(* Logix 5000 project; controller PLC_MCC1300_75F1 vendor 1 type 14 code 166 rev 32.11; software revision 32.04; part 68 of 83 *)
(* tags used below, declared in another part *)
   CM_AreaStackerToLine_JS1_Sync : CM_AreaStackerToLine;
   CM_ConveyorStackerToLine_JS1_Sync : CM_ConveyorStackerToLine;
   CM_DATA_Z410_Rx_Sync : UDT_PlateData_Convoy;
   CM_DATA_Z410_Tx : UDT_PlateData_Convoy;
   CM_DATA_Z410_Tx_PH : DINT;
   CM_LineToAreaStacker_JS1 : CM_LineToAreaStacker;
   CM_LineToConveyorStacker_JS1 : CM_LineToConveyorStacker;
   CM_LineToConveyorStacker_JS2 : CM_LineToConveyorStacker;
   GP_AccessArea_M311S_STC : GP_AccessArea_STC;
   GP_ConvertDataFromStacker : GP_ConvertDataFromStacker;
   GP_ConvertDataToStacker : GP_ConvertDataToStacker;
   Gp_SpaceConvUtilities_V1 : GP_SpaceConvUtilities_V1;
   M311 : MAC_Conveyor;
   M311_SpaceConv_Utilities : SpaceConv_Utilities;
   M316 : MAC_Conveyor;
   M316_SpaceConv_Utilities : SpaceConv_Utilities;
   M317 : MAC_Conveyor_Single;
   M317_Data : UDT_Convoy_SL;
   M317_dTractionRecovery_M3 : DINT;
   M317_dTractionRecovery_M4 : DINT;
   M317_HMR : MAC_Conveyor_HMR;
   M317_HMW : MAC_Conveyor_HMW;
   M317_M3_DR_IN_MAM : MOTION_INSTRUCTION;
   M317_M3_DR_IN_MRP : MOTION_INSTRUCTION;
   M317_SpaceConv_Utilities : SpaceConv_Utilities;
   M317_xEnableTractionRecovering : BOOL;
   M317_xLateralTractionRecovered : BOOL;
   M317_xSendCulletReqActive : BOOL;
   O : INT[128];
   TMP_CenterLites : BOOL;
   TMP_d : DINT;
   TMP_dDecelerationPositionEndConveyor : DINT;
   TMP_DistanceLateralSquaringToCenter : DINT;
   TMP_dOffsetLoadUnload_cmm : DINT;
   TMP_SendToCullet : BOOL;
   TMP_SquaringPosition : DINT;
   TMP_xConveyorOfStartCleaning : BOOL;
   TMP_xCulletPresent : BOOL;
   TMP_xLiteThisDestPresent : BOOL;
   xAlwaysOFF : BOOL;
   xAlwaysON : BOOL;
   xDebugOFF : BOOL;
   Z402 : MAC_Zone;
   Z402_HMR : MAC_Zone_HMR;
   Z402S_INPUT_xSafetyAreaPopup : BOOL;
(* MainProgram, continued *)

   // Calculation Space for Wait Stop Next Conveyor
   39: CPT(TMP_dDecelerationPositionEndConveyor,M317_SpaceConv_Utilities.CONST_dConveyorLength_cmm - M317.AUX_dAccSpace_cmm + 1000);
   // Wait stop next Machine
   40: XIO(M317.PH_x.8)GEQ(M317_SpaceConv_Utilities.O_dHeadPosition_cmm,TMP_dDecelerationPositionEndConveyor)OTE(M317.ST_xWaitStopNextMachine);
   // Set Wait Machine Stop
   41: [XIC(M317.PH_x.7) [XIO(xAlwaysOFF) ,XIC(M317.ST_xWaitStopNextMachine) [XIC(M311_SpaceConv_Utilities.O_xRampInProgress) ,XIO(M311_SpaceConv_Utilities.ST_xFeedbackRotation) ] ] ,XIC(M317.PH_x.0) NEQ(Z402_HMR.dLineSpeed_mm_min,M317.AUX_dReqSpeed_mm_min) ]OTL(M317.ST_xWaitMachineStop);
   // Reset Wait Machine Stop
   42: XIO(M317_SpaceConv_Utilities.ST_xFeedbackRotation)[XIO(M317_SpaceConv_Utilities.ST_xFeedbackRotation) ,XIO(M317.ST_xWaitStopNextMachine) ]EQU(Z402_HMR.dLineSpeed_mm_min,M317.AUX_dReqSpeed_mm_min)OTU(M317.ST_xWaitMachineStop);
   // Request send plate_data to stacker
   43: XIO(M317_xSendCulletReqActive)XIO(xDebugOFF)XIO(M317.PH_x.8)XIO(M317.PH_x.15)XIO(xDebugOFF)XIC(Z402.ST_xConditionOkPhaseAdvancement)XIC(M317.ST_xPlatePresence)XIC(M317.ST_xIdPlatePresence)XIC(M317.ST_xOutputEnable)XIO(M317.ST_xWaitMachineStop)XIO(M317_Data.rgtCap[0].rgxRequest.0)XIO(M317_Data.rgtCap[0].rgxRequest.1)XIO(M317_Data.rgtCap[0].rgxRequest.2)XIC(TMP_xLiteThisDestPresent)[GP_ConvertDataToStacker(GP_ConvertDataToStacker,M317_Data,CM_DATA_Z410_Tx) ,XIO(CM_DATA_Z410_Tx_PH.6) XIO(CM_LineToConveyorStacker_JS2.xRequestForUnload) OTL(CM_DATA_Z410_Tx_PH.0) ,OTE(CM_LineToConveyorStacker_JS2.xRequestForUnload) ];
   44: XIC(CM_LineToConveyorStacker_JS1.xRequestForUnload)XIC(CM_DATA_Z410_Tx_PH.6)TON(M317.TmON[2],?,?)XIC(M317.TmON[2].DN)OTU(CM_DATA_Z410_Tx_PH.6)OTL(CM_DATA_Z410_Tx_PH.0);
   // Phase of unload
   45: XIO(M317_xSendCulletReqActive)XIC(Z402.ST_xConditionOkPhaseAdvancement)XIC(M317.ST_xPlatePresence)XIC(M317.ST_xIdPlatePresence)XIC(M317.ST_xOutputEnable)XIO(M317.ST_xWaitMachineStop)XIO(M317.PH_x.8)XIO(M317_Data.rgtCap[0].rgxRequest.0)XIO(M317_Data.rgtCap[0].rgxRequest.1)XIO(M317_Data.rgtCap[0].rgxRequest.2)XIC(M317.INPUT_xLowPositionSquaring_1)XIC(M317.INPUT_xLowPositionPopup_1)XIC(M317.INPUT_xLowPositionPopup_2)XIC(TMP_xLiteThisDestPresent)XIC(CM_ConveyorStackerToLine_JS1_Sync.xInitialContionOk)XIO(CM_DATA_Z410_Tx_PH.0)XIO(CM_DATA_Z410_Tx_PH.3)EQU(CM_LineToAreaStacker_JS1.dMsgDataSync,CM_AreaStackerToLine_JS1_Sync.dMsgDataSyncFdbk)EQU(CM_DATA_Z410_Tx.dSyncHead,CM_AreaStackerToLine_JS1_Sync.dMsgDataSyncFdbk)[OTE(M317.ST_xWaitReadyToMove) ,[XIC(M317.ST_xAxleReadyToMoveDelayed) ,XIC(xAlwaysON) ] [OTE(M317.OS_xUnload_FW) ,OTL(M317.PH_x.8) ,MOV(M317_Data.dLength_cmm,M317_SpaceConv_Utilities.CONF_MD4_MD6_dLength_cmm) GP_SpaceConvUtilities_V1(Gp_SpaceConvUtilities_V1,M317_SpaceConv_Utilities,M316_SpaceConv_Utilities,M317_SpaceConv_Utilities,6) ,FLL(0,M317_Data,1) ] ];
   // Phase of end unload
   46: XIC(M317.PH_x.8)[GEQ(M317_SpaceConv_Utilities.O_dTailPosition_cmm,M317.AUX_dPresetStopUnload_cmm) ,XIO(M317_SpaceConv_Utilities.ST_xFeedbackRotation) GEQ(M317_SpaceConv_Utilities.O_dTailPosition_cmm,M317_SpaceConv_Utilities.CONST_dConveyorLength_cmm) ][OTE(M317.PH_x.15) ,OTU(M317.PH_x.8) ,OTU(M317.ST_xPlatePresence) ];
   // Frontal squaring management
   // -
   // -
   47: NOP();
   // Frontal squaring phase
   48: XIC(Z402.ST_xConditionOkPhaseAdvancement)XIC(M317.ST_xPlatePresence)XIC(M317.ST_xIdPlatePresence)XIC(M317.ST_xOutputEnable)XIC(M317_Data.rgtCap[0].rgxRequest.0)[XIO(M317.ST_xPhasesInProgress) ,XIC(M317.PH_x.7) ]XIO(M317.INPUT_xSyncroPhotocell_1)XIO(M317.INPUT_xSyncroPhotocell_2)OTL(M317.PH_x.4);
   // Position squaring set
   49: XIC(M317.PH_x.4)GEQ(M317_SpaceConv_Utilities.O_dHeadPosition_cmm,TMP_SquaringPosition)CPT(M317_SpaceConv_Utilities.CONF_MD2_MD3_dPrstPos_cmm,TMP_SquaringPosition)GP_SpaceConvUtilities_V1(Gp_SpaceConvUtilities_V1,M317_SpaceConv_Utilities,M316_SpaceConv_Utilities,M317_SpaceConv_Utilities,2);
   // End Frontal squaring phase
   50: XIC(M317.PH_x.4)[[GEQ(M317_SpaceConv_Utilities.O_dHeadPosition_cmm,TMP_SquaringPosition) [XIC(M317.INPUT_xSquaringPhotocell_1) ,XIC(M317.INPUT_xSquaringPhotocell_2) ] ,XIC(M317.INPUT_xSquaringPhotocell_1) ,XIC(M317.INPUT_xSquaringPhotocell_2) ] ,XIC(M317.ST_xPhaseError) ][MOV(M317_HMW.dParam_5_ms,M317.tmON_AuxFunction5.PRE) TON(M317.tmON_AuxFunction5,?,?) ,[XIC(M317.tmON_AuxFunction5.DN) ,XIC(M317.ST_xPhaseError) ] [OTU(M317.PH_x.4) ,OTE(M317.PH_x.5) ,OTU(M317_Data.rgtCap[0].rgxRequest.0) ,XIO(M317.ST_xPhaseError) OTL(M317_Data.rgtCap[0].rgxDone.0) ] ];
   // Popup management
   // -
   // -
   51: NOP();
   // Phase of Rise popup
   52: XIC(Z402.ST_xConditionOkPhaseAdvancement)XIC(M317.ST_xPlatePresence)XIC(M317.ST_xIdPlatePresence)XIC(M317.ST_xOutputEnable)XIO(M317.ST_xPhasesInProgress)XIO(M317.INPUT_xHighPositionPopup_1)XIO(TMP_xCulletPresent)[XIC(M317_Data.rgtCap[0].rgxRequest.1) [XIC(M317_xEnableTractionRecovering) XIC(M317_xLateralTractionRecovered) ,XIO(M317_xEnableTractionRecovering) ] ,XIC(M317_Data.rgtCap[0].rgxRequest.2) [XIC(M317_xEnableTractionRecovering) XIC(M317_xLateralTractionRecovered) ,XIO(M317_xEnableTractionRecovering) ] ]OTL(M317.PH_x.16);
   // Phase of End rise popup
   53: XIC(M317.PH_x.16)XIC(M317.INPUT_xHighPositionPopup_1)XIC(M317.INPUT_xHighPositionPopup_2)[OTU(M317.PH_x.16) ,OTE(M317.PH_x.19) ];
   // Phase of descent popup
   54: XIC(Z402.ST_xConditionOkPhaseAdvancement)XIC(M317.ST_xOutputEnable)XIO(M317.ST_xPhasesInProgress)XIO(M317.INPUT_xLowPositionPopup_1)XIO(M317.INPUT_xLowPositionPopup_2)XIO(M317_Data.rgtCap[0].rgxRequest.1)XIO(M317_Data.rgtCap[0].rgxRequest.2)XIO(M317_Data.rgtCap[0].rgxRequest.3)OTL(M317.PH_x.20);
   // Phase of end descent popup
   55: XIC(M317.PH_x.20)XIC(M317.INPUT_xLowPositionPopup_1)XIC(M317.INPUT_xLowPositionPopup_2)[OTU(M317.PH_x.20) ,OTE(M317.PH_x.23) ,XIO(xAlwaysOFF) OTU(M317_xLateralTractionRecovered) ];
   // Lateral squaring management
   // -
   // -
   56: NOP();
   57: XIC(Z402.ST_xConditionOkPhaseAdvancement)XIC(M317.ST_xPlatePresence)XIC(M317.ST_xOutputEnable)XIO(M317.ST_xPhasesInProgress)XIC(M317.INPUT_xHighPositionPopup_1)XIC(M317_Data.rgtCap[0].rgxRequest.1)OTL(M317.PH_x.28);
   58: XIC(M317.PH_x.28)[NEQ(M317_Data.rgtCap[0].rgtLite[0].dID,0) MOV(M317_HMW.dParam_7_ms,M317.tmON_AuxFunction2.PRE) XIC(M317.INPUT_xSquaringPhotocell_3) TON(M317.tmON_AuxFunction2,?,?) ,NEQ(M317_Data.rgtCap[0].rgtLite[1].dID,0) MOV(M317_HMW.dParam_7_ms,M317.tmON_AuxFunction3.PRE) XIC(M317.INPUT_xSquaringPhotocell_4) TON(M317.tmON_AuxFunction3,?,?) ];
   59: XIC(M317.PH_x.28)[[XIC(M317.tmON_AuxFunction2.DN) ,EQU(M317_Data.rgtCap[0].rgtLite[0].dID,0) ] [XIC(M317.tmON_AuxFunction3.DN) ,EQU(M317_Data.rgtCap[0].rgtLite[1].dID,0) ] ,XIC(M317.ST_xPhaseError) ][OTU(M317.PH_x.28) ,OTE(M317.PH_x.29) ,XIO(M317.ST_xPhaseError) [NEQ(M317_Data.rgtCap[0].rgtLite[0].dID,0) CPT(M317_Data.rgtCap[0].rgtLite[0].dBarycenter_cmm,M317_Data.rgtCap[0].rgtLite[0].dWidth_cmm / 2 - TMP_DistanceLateralSquaringToCenter) ,NEQ(M317_Data.rgtCap[0].rgtLite[1].dID,0) CPT(M317_Data.rgtCap[0].rgtLite[1].dBarycenter_cmm,TMP_DistanceLateralSquaringToCenter - M317_Data.rgtCap[0].rgtLite[1].dWidth_cmm / 2) ] ,OTU(M317_Data.rgtCap[0].rgxRequest.1) ,XIO(M317.ST_xPhaseError) OTL(M317_Data.rgtCap[0].rgxDone.1) ];
   // Adjust Y position management
   // -
   // -
   60: NOP();
   61: XIO(M317_xSendCulletReqActive)XIC(Z402.ST_xConditionOkPhaseAdvancement)XIC(M317.ST_xPlatePresence)XIC(M317.ST_xOutputEnable)XIO(M317.ST_xPhasesInProgress)[XIC(M317_Data.rgtCap[0].rgxRequest.2) ,XIC(M317_xEnableTractionRecovering) XIC(M317_Data.rgtCap[0].rgxRequest.1) ][XIC(M317_Data.rgtCap[0].rgxRequest.2) [XIO(M317_xEnableTractionRecovering) XIC(M317.INPUT_xHighPositionPopup_1) XIC(M317.INPUT_xHighPositionPopup_2) ,XIC(M317_xEnableTractionRecovering) XIC(M317_xLateralTractionRecovered) ] ,[XIC(M317_Data.rgtCap[0].rgxRequest.1) ,XIC(M317_Data.rgtCap[0].rgxRequest.2) ] XIC(M317_xEnableTractionRecovering) XIO(M317_xLateralTractionRecovered) XIC(M317.INPUT_xLowPositionPopup_1) XIC(M317.INPUT_xLowPositionPopup_2) ]XIO(M317.INPUT_xDriveFeedback_M3)XIO(M317.INPUT_xDriveFeedback_M4)OTL(M317.PH_x.24);
   // Target positioning M3 & M4
   62: XIC(M317.PH_x.24)XIC(TMP_CenterLites)[CPT(M317.AUX_dAbsPosTarget_M3_cmm,- ((M317_Data.rgtCap[0].rgtLite[0].dBarycenter_cmm + M317_Data.rgtCap[0].rgtLite[1].dBarycenter_cmm) / 2)) ,MOV(M317.AUX_dAbsPosTarget_M3_cmm,M317.AUX_dAbsPosTarget_M4_cmm) ];
   63: XIC(M317.PH_x.24)[XIC(M317_M3_DR_IN_MRP.EN) XIC(M317_M3_DR_IN_MRP.DN) ,XIC(M317.ST_xPhaseError) ][OTU(M317.PH_x.24) ,[XIC(M317_xEnableTractionRecovering) XIC(M317_xLateralTractionRecovered) ,XIO(M317_xEnableTractionRecovering) ] XIC(M317.INPUT_xHighPositionPopup_1) XIC(M317.INPUT_xHighPositionPopup_2) OTL(M317.PH_x.26) ,XIC(M317_xEnableTractionRecovering) XIO(M317_xLateralTractionRecovered) [OTL(M317.PH_x.30) ,[GRT(M317.AUX_dAbsPosTarget_M3_cmm,0) MOV(1500,M317_dTractionRecovery_M3) ,LES(M317.AUX_dAbsPosTarget_M3_cmm,0) MOV(-1500,M317_dTractionRecovery_M3) ,GRT(M317.AUX_dAbsPosTarget_M4_cmm,0) MOV(1500,M317_dTractionRecovery_M4) ,LES(M317.AUX_dAbsPosTarget_M4_cmm,0) MOV(-1500,M317_dTractionRecovery_M4) ] ] ];
   64: XIC(M317.PH_x.30)[XIC(M317.OUTPUT_xPositioning_M3) XIC(M317.OUTPUT_xPositioning_M4) XIC(M317_M3_DR_IN_MAM.EN) XIC(M317_M3_DR_IN_MAM.PC) ,XIC(M317.ST_xPhaseError) ][OTU(M317.PH_x.30) ,OTE(M317.PH_x.31) ,XIO(M317.ST_xPhaseError) OTL(M317_xLateralTractionRecovered) ];
   65: XIC(M317.PH_x.26)[XIC(M317.OUTPUT_xPositioning_M3) XIC(M317.OUTPUT_xPositioning_M4) XIC(M317_M3_DR_IN_MAM.EN) XIC(M317_M3_DR_IN_MAM.PC) ,XIC(M317.ST_xPhaseError) ][OTU(M317.PH_x.26) ,OTE(M317.PH_x.27) ,OTU(M317_Data.rgtCap[0].rgxRequest.2) ,XIO(M317.ST_xPhaseError) OTL(M317_Data.rgtCap[0].rgxDone.2) ];
   66: XIC(M317.PH_x.27)XIO(M317.ST_xPhaseError)[NEQ(M317_Data.rgtCap[0].rgtLite[0].dID,0) ADD(M317_Data.rgtCap[0].rgtLite[0].dBarycenter_cmm,M317.AUX_dAbsPosTarget_M3_cmm,M317_Data.rgtCap[0].rgtLite[0].dBarycenter_cmm) ,NEQ(M317_Data.rgtCap[0].rgtLite[1].dID,0) ADD(M317_Data.rgtCap[0].rgtLite[1].dBarycenter_cmm,M317.AUX_dAbsPosTarget_M4_cmm,M317_Data.rgtCap[0].rgtLite[1].dBarycenter_cmm) ];
   // Phase of load (from M409) NEGATIVE
   67: XIC(CM_ConveyorStackerToLine_JS1_Sync.xRequestReturnInLine)XIC(CM_ConveyorStackerToLine_JS1_Sync.xRotationForUnload)[NEQ(CM_DATA_Z410_Rx_Sync.tLite[0].dID,0) ,NEQ(CM_DATA_Z410_Rx_Sync.tLite[1].dID,0) ]XIO(M317.ST_xPhasesInProgress)[OTL(M317.PH_x.10) ,OTU(M317_SpaceConv_Utilities.O_xPlateSynchronized) ,OTU(M317.ST_xDisableLoadUnloadOnStop) ,OTE(M317.OS_xLoad_BW) ,GP_ConvertDataFromStacker(GP_ConvertDataFromStacker,CM_DATA_Z410_Rx_Sync,M317_Data) FLL(0,CM_DATA_Z410_Rx_Sync,1) ,GP_SpaceConvUtilities_V1(Gp_SpaceConvUtilities_V1,M317_SpaceConv_Utilities,M316_SpaceConv_Utilities,M317_SpaceConv_Utilities,15) ,MOV(-135000,M317_SpaceConv_Utilities.CONF_MD2_MD3_dPrstPos_cmm) GP_SpaceConvUtilities_V1(Gp_SpaceConvUtilities_V1,M317_SpaceConv_Utilities,M316_SpaceConv_Utilities,M317_SpaceConv_Utilities,2) ];
   // Syncro  -  Space Convoy utilities MOD 4
   // verificare se esiste la sincro quando si carica in backward
   68: GRT(M317_SpaceConv_Utilities.CONST_dSyncMode,0)[XIC(M317.PH_x.10) XIO(M317.PH_x.12) ,XIC(M317.PH_x.10) XIC(M317.PH_x.12) ADD(M317_SpaceConv_Utilities.CONST_dSyncroPhPosition_cmm,TMP_dOffsetLoadUnload_cmm,TMP_d) GRT(M317_SpaceConv_Utilities.O_dTailPosition_cmm,TMP_d) ][MOV(M317_Data.dLength_cmm,M317_SpaceConv_Utilities.CONF_MD4_MD6_dLength_cmm) ,GP_SpaceConvUtilities_V1(Gp_SpaceConvUtilities_V1,M317_SpaceConv_Utilities,M316_SpaceConv_Utilities,M317_SpaceConv_Utilities,4) ];
   // End load Phase (from M409) NEGATIVE
   69: XIC(M317.PH_x.10)[GRT(M317_SpaceConv_Utilities.O_dHeadPosition_cmm,M317.AUX_dPresetStopLoad_cmm) ,CPT(TMP_d,M317_SpaceConv_Utilities.CONST_dConveyorLength_cmm/2 + M317_Data.dLength_cmm / 2) GRT(M317_SpaceConv_Utilities.O_dHeadPosition_cmm,TMP_d) ][OTE(M317.PH_x.11) ,OTU(M317.PH_x.10) ,OTL(M317.ST_xPlatePresence) ];
   // Phase of unload (to M316) NEGATIVE
   70: XIC(Z402.ST_xConditionOkPhaseAdvancement)XIC(M317.ST_xPlatePresence)XIC(M317.ST_xIdPlatePresence)XIC(M317.ST_xOutputEnable)XIO(M317.ST_xWaitMachineStop)XIO(M317.PH_x.12)XIO(TMP_xLiteThisDestPresent)XIO(M317.ST_xPhasesInProgress)XIC(M317.INPUT_xLowPositionPopup_1)XIC(M317.INPUT_xLowPositionPopup_2)XIO(M317.ST_xVirtualDoorEnabled)[XIC(M311.ST_xInitialConditionOK_BW) XIO(M317.ST_xVirtualDoorEnabled) [XIC(M317.ST_xAxleReadyToMoveDelayed) ,XIC(xAlwaysON) ] [OTE(M317.OS_xUnload_BW) ,OTL(M317.PH_x.12) ,MOV(M317_Data.dLength_cmm,M317_SpaceConv_Utilities.CONF_MD4_MD6_dLength_cmm) GP_SpaceConvUtilities_V1(Gp_SpaceConvUtilities_V1,M317_SpaceConv_Utilities,M316_SpaceConv_Utilities,M317_SpaceConv_Utilities,16) ] ,OTE(M317.ST_xAux1) ];
   // Phase of end unload (to M316) NEGATIVE
   71: XIC(M317.PH_x.12)[GEQ(M317_SpaceConv_Utilities.O_dTailPosition_cmm,M317.AUX_dPresetStopUnload_cmm) ,XIO(M317_SpaceConv_Utilities.ST_xFeedbackRotation) GEQ(M317_SpaceConv_Utilities.O_dTailPosition_cmm,M317_SpaceConv_Utilities.CONST_dConveyorLength_cmm) ][OTE(M317.PH_x.13) ,OTU(M317.PH_x.12) ,OTU(M317.ST_xPlatePresence) ];
   // Redestination lites
   // -
   // -
   72: [XIC(M317.ST_xPhaseError) [XIC(M317.PH_x.7) XIC(M317_Data.tFlag.tConveyor.xReqStop) ,XIC(M317.PH_x.5) ,XIC(M317.PH_x.29) ,XIC(M317.PH_x.27) ] ,[XIC(CM_AreaStackerToLine_JS1_Sync.xSB_SendToCullet) ,XIC(CM_AreaStackerToLine_JS1_Sync.xSB_DestinationChange) ] ,[XIC(CM_ConveyorStackerToLine_JS1_Sync.xRequestReturnInLine) ,XIO(CM_AreaStackerToLine_JS1_Sync.xStackerInUnloaderMode) ] XIC(TMP_xLiteThisDestPresent) ,XIC(M317_xSendCulletReqActive) XIO(M317.ST_xPhasesInProgress) ]OTL(TMP_SendToCullet)OTU(M317.ST_xPhaseError);
   // Phase in progress
   73: NEQ(M317.PH_x,0)OTE(M317.ST_xPhasesInProgress);
   // #####_CLEANING_#####
   74: NOP();
   // Cleaning Reset
   75: XIC(M317.ST_xCleaningAccepted)[XIC(Z402.ST_xCleaningAccepted) ,XIO(TMP_xConveyorOfStartCleaning) ][XIC(M317.ST_xIdPlatePresence) OTL(TMP_SendToCullet) FLL(0,M317_Data,1) ,MOV(0,M317.PH_x) OTU(M317.ST_xPlatePresence) ];
   // Initial condition OK
   76: XIC(Z402.ST_xConditionOkPhaseAdvancement)XIC(M317.ST_xOutputEnable)XIO(M317_HMW.xEnableDisableManualCommand)XIO(M317.ST_xReqCleaning)XIO(M317.ST_xCleaningAccepted)XIO(M317.ST_xStopNextCycleFault)XIO(M317.ST_xVirtualDoorEnabled)XIO(M317.PH_x.0)[XIO(M317.ST_xPhasesInProgress) XIO(M317.ST_xPlatePresence) ,XIC(M317.ST_xCycleLoadUnload) XIC(M317.PH_x.8) XIC(M317.OUTPUT_xRun_M1) GRT(M317_SpaceConv_Utilities.O_dTailPosition_cmm,M317_SpaceConv_Utilities.O_dPresetLoadUnload_cmm) XIO(M317.ST_xIdPlatePresence) ]XIC(M317.INPUT_xLowPositionPopup_1)XIC(M317.INPUT_xLowPositionPopup_2)XIO(CM_ConveyorStackerToLine_JS1_Sync.xRequestReturnInLine)XIO(GP_AccessArea_M311S_STC.ST_xAccessRequest)XIO(GP_AccessArea_M311S_STC.ST_xAccessAccepted)XIC(Z402S_INPUT_xSafetyAreaPopup)OTE(M317.ST_xInitialConditionOK);
   // Initial condition OK (M409)
   77: XIC(Z402.ST_xConditionOkPhaseAdvancement)XIC(M317.ST_xOutputEnable)XIO(M317_HMW.xEnableDisableManualCommand)XIO(M317.ST_xReqCleaning)XIO(M317.ST_xCleaningAccepted)XIO(M317.ST_xStopNextCycleFault)XIC(M317.INPUT_xLowPositionPopup_1)XIC(M317.INPUT_xLowPositionPopup_2)XIO(M317.INPUT_xHighPositionSquaring_1)XIO(M317.ST_xPhasesInProgress)XIO(M317.ST_xPlatePresence)XIC(CM_ConveyorStackerToLine_JS1_Sync.xRequestReturnInLine)XIO(GP_AccessArea_M311S_STC.ST_xAccessRequest)XIO(GP_AccessArea_M311S_STC.ST_xAccessAccepted)XIC(Z402S_INPUT_xSafetyAreaPopup)OTE(M317.ST_xInitialConditionOK_BW);
   // #####_HMI_STATUSES_#####
   78: NOP();
   // PhotocelPresence {x|x|x|x|O}
   79: XIC(M317.INPUT_xSyncroPhotocell_1)OTE(M317_HMR.xSensorPresence5);
   // PhotocelPresence {x|x|x|x|O}
   80: XIC(M317.INPUT_xSyncroPhotocell_2)OTE(M317_HMR.xSensorPresence6);
   // Frontal squaring photocell {x|x|x|x|O}
   81: XIC(M317.INPUT_xSquaringPhotocell_1)OTE(M317_HMR.xSensorPresence3);
   // Right squaring photocell {x|x|x|x|O}
   82: XIC(M317.INPUT_xSquaringPhotocell_2)OTE(M317_HMR.xSensorPresence4);
   // Left squaring photocell {x|x|x|x|O}
   83: XIC(M317.INPUT_xSquaringPhotocell_3)OTE(M317_HMR.xSensorPresence1);
   // Left squaring photocell {x|x|x|x|O}
   84: XIC(M317.INPUT_xSquaringPhotocell_4)OTE(M317_HMR.xSensorPresence2);
   // High position popup {x|x|x|x|O}
   85: XIC(M317.INPUT_xHighPositionPopup_1)OTE(M317_HMR.xHighPositionPopup1);
   // High position popup {x|x|x|x|O}
   86: XIC(M317.INPUT_xHighPositionPopup_2)OTE(M317_HMR.xHighPositionPopup2);
   // Low position popup {x|x|x|x|O}
   87: XIC(M317.INPUT_xLowPositionPopup_1)OTE(M317_HMR.xLowPositionPopup1);
   // Low position popup {x|x|x|x|O}
   88: XIC(M317.INPUT_xLowPositionPopup_2)OTE(M317_HMR.xLowPositionPopup2);
   // High position frontal squaring {x|x|x|x|O}
   89: XIC(M317.INPUT_xHighPositionSquaring_1)OTE(M317_HMR.xHighPositionSquaring1)OTE(M317_HMR.xHighPositionSquaring2);
   // Low position frontal squaring {x|x|x|x|O}
   90: XIC(M317.INPUT_xLowPositionSquaring_1)OTE(M317_HMR.xLowPositionSquaring1)OTE(M317_HMR.xLowPositionSquaring2);
   // Manual Mode Enable {x|x|x|x|O}
   91: XIC(M317.ST_xManualMode)OTE(M317_HMR.xManualCommandEnabled);
   // Command forward M1
   92: XIC(M317.ST_xManualMode)XIC(M317_HMW.rgxMan.0)XIC(M317.OUTPUT_xRun_M1)OTE(M317_HMR.rgxMan.0);
   // Command backward M1
   93: XIC(M317.ST_xManualMode)XIC(M317_HMW.rgxMan.1)XIC(M317.OUTPUT_xReverse_M1)OTE(M317_HMR.rgxMan.1);
   // Command forward M2
   94: XIC(M317.ST_xManualMode)XIC(M317_HMW.rgxMan.2)XIC(M317.OUTPUT_xRun_M2)OTE(M317_HMR.rgxMan.2);
   // Command backward M2
   95: XIC(M317.ST_xManualMode)XIC(M317_HMW.rgxMan.3)XIC(M317.OUTPUT_xReverse_M2)OTE(M317_HMR.rgxMan.3);
   // Command forward M3
   96: XIC(M317.ST_xManualMode)XIC(M317_HMW.rgxMan.4)XIC(M317.OUTPUT_xRun_M3)OTE(M317_HMR.rgxMan.4);
   // Command backward M3
   97: XIC(M317.ST_xManualMode)XIC(M317_HMW.rgxMan.5)XIC(M317.OUTPUT_xReverse_M3)OTE(M317_HMR.rgxMan.5);
   // Command forward M4
   98: XIC(M317.ST_xManualMode)XIC(M317_HMW.rgxMan.6)XIC(M317.OUTPUT_xRun_M4)OTE(M317_HMR.rgxMan.6);
   // Command backward M4
   99: XIC(M317.ST_xManualMode)XIC(M317_HMW.rgxMan.7)XIC(M317.OUTPUT_xReverse_M4)OTE(M317_HMR.rgxMan.7);
   // Command rise frontal squaring
   100: XIC(M317.ST_xManualMode)XIC(M317_HMW.rgxMan.10)XIC(M317.OUTPUT_xRiseSquaring_1)OTE(M317_HMR.rgxMan.10);
   // Command descent frontal squaring
   101: XIC(M317.ST_xManualMode)XIC(M317_HMW.rgxMan.11)XIC(M317.OUTPUT_xDescentSquaring_1)OTE(M317_HMR.rgxMan.11);
   // Command rise frontal squaring
   102: XIC(M317.ST_xManualMode)XIC(M317_HMW.rgxMan.16)XIC(M317.OUTPUT_xRiseSquaring_1)OTE(M317_HMR.rgxMan.16);
